(* Logix 5000 project; controller WED2413001_BI600_AB vendor 1 type 14 code 192 rev 35.11; software revision 35.01 *) (continued)
   TRANSITION Tran_008 FROM R00STARTING TO R00EXECUTE
      := EXECUTING
   END_TRANSITION
   STEP R00EXECUTE:
      ACTION Action_008 (N):
         Machine_State:=6;
      END_ACTION
   END_STEP
   TRANSITION Tran_011 FROM R00EXECUTE TO R00STOPPING
      := 
         STOP_CMD
   END_TRANSITION
   TRANSITION Tran_012 FROM R00EXECUTE TO R00COMPLETING
      := PRODUCTION_CNT
   END_TRANSITION
   TRANSITION Tran_009 FROM R00EXECUTE TO R00SUSPENDING
      := SUSPEND_CMD
   END_TRANSITION
   TRANSITION Tran_010 FROM R00EXECUTE TO R00HOLDING
      := HOLD_CMD
   END_TRANSITION
   STEP R00STOPPING:
      ACTION Action_009 (N):
         Machine_State:=7;
      END_ACTION
   END_STEP
   STEP R00COMPLETING:
      ACTION Action_010 (N):
         Machine_State:=16;
      END_ACTION
   END_STEP
   STEP R00SUSPENDING:
      ACTION Action_011 (N):
         Machine_State:=13;
      END_ACTION
   END_STEP
   STEP R00HOLDING:
      ACTION Action_012 (N):
         Machine_State:=10;
      END_ACTION
   END_STEP
   TRANSITION Tran_013 FROM R00STOPPING TO R00STOPPED
      := 1
   END_TRANSITION
   TRANSITION Tran_014 FROM R00COMPLETING TO R00COMPLETE
      := 1
   END_TRANSITION
   TRANSITION Tran_015 FROM R00SUSPENDING TO R00SUSPENDED
      := SUSPEND_CMD
   END_TRANSITION
   TRANSITION Tran_016 FROM R00HOLDING TO R00HELD
      := HOLD_CMD
   END_TRANSITION
   STEP R00COMPLETE:
      ACTION Action_015 (N):
         Machine_State:=17;
      END_ACTION
   END_STEP
   STEP R00SUSPENDED:
      ACTION Action_014 (N):
         Machine_State:=5;
      END_ACTION
   END_STEP
   STEP R00HELD:
      ACTION Action_013 (N):
         Machine_State:=11;
      END_ACTION
   END_STEP
   TRANSITION Tran_017 FROM R00COMPLETE TO R00RESETING
      := 1
   END_TRANSITION
   TRANSITION Tran_018 FROM R00SUSPENDED TO R00UNSUSPENDED
      := SUSPEND_CMD
   END_TRANSITION
   TRANSITION Tran_019 FROM R00HELD TO R00UNHOLDING
      := RESUME_CMD
   END_TRANSITION
   STEP R00UNSUSPENDED:
      ACTION Action_016 (N):
         Machine_State:=14;
      END_ACTION
   END_STEP
   STEP R00UNHOLDING:
      ACTION Action_017 (N):
         Machine_State:=12;
      END_ACTION
   END_STEP
   TRANSITION Tran_020 FROM R00UNSUSPENDED TO R00EXECUTE
      := 1
   END_TRANSITION
   TRANSITION Tran_021 FROM R00UNHOLDING TO R00EXECUTE
      := 1
   END_TRANSITION
END_ROUTINE

ROUTINE R00_Main   (* ladder *)
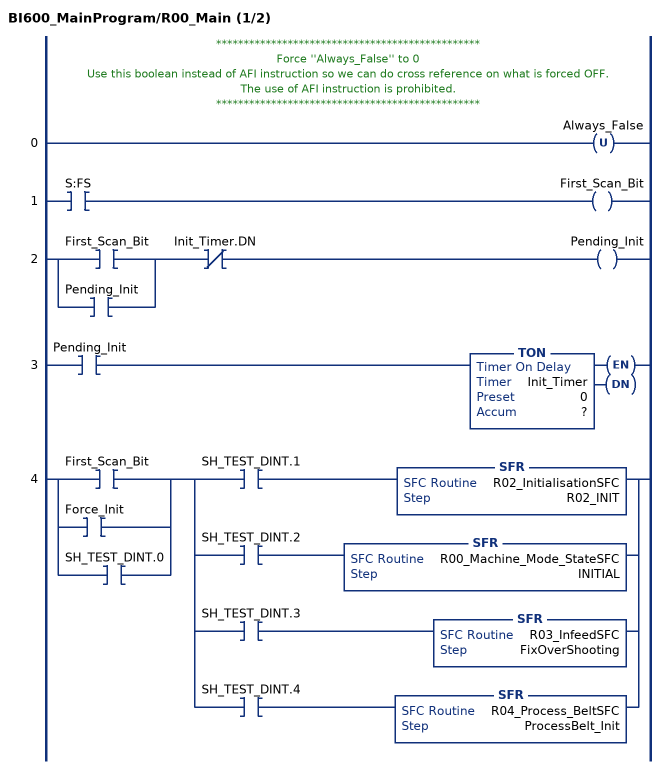
   // ************************************************
   // Force ''Always_False'' to 0
   // Use this boolean instead of AFI instruction so we can do cross reference on what is forced OFF.
   // The use of AFI instruction is prohibited.
   // ************************************************
   0: OTU(Always_False);
   1: XIC(S:FS)OTE(First_Scan_Bit);
   2: [XIC(First_Scan_Bit) ,XIC(Pending_Init) ]XIO(Init_Timer.DN)OTE(Pending_Init);
   3: XIC(Pending_Init)TON(Init_Timer,?,?);
   4: [XIC(First_Scan_Bit) ,XIC(Force_Init) ,XIC(SH_TEST_DINT.0) ][XIC(SH_TEST_DINT.1) SFR(R02_InitialisationSFC,R02_INIT) ,XIC(SH_TEST_DINT.2) SFR(R00_Machine_Mode_StateSFC,INITIAL) ,XIC(SH_TEST_DINT.3) SFR(R03_InfeedSFC,FixOverShooting) ,XIC(SH_TEST_DINT.4) SFR(R04_Process_BeltSFC,ProcessBelt_Init) ];
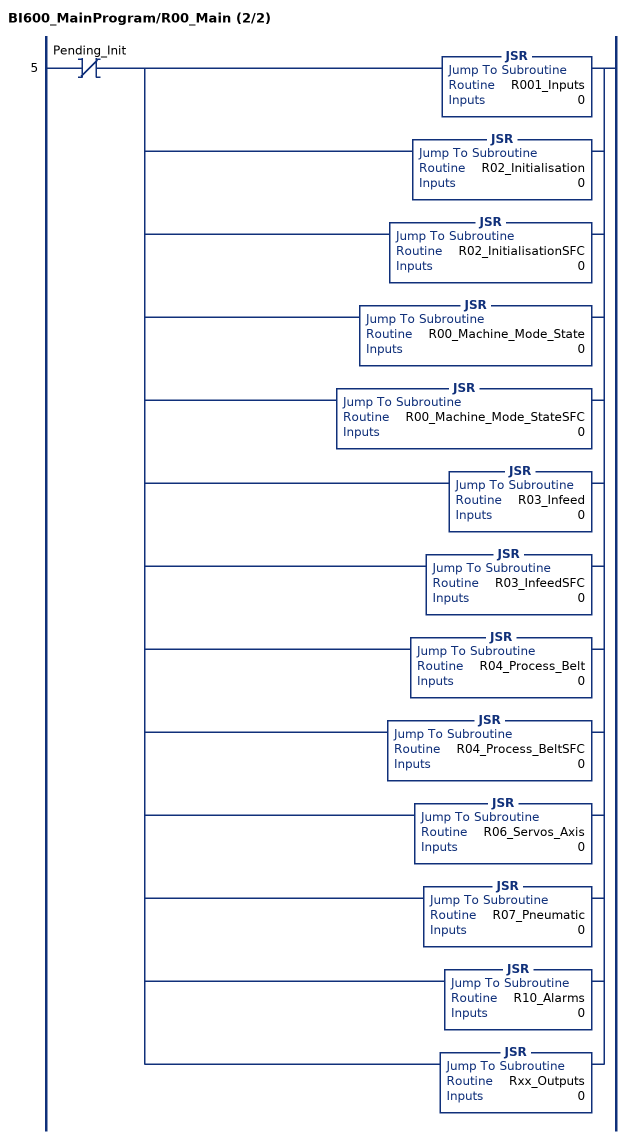
   5: XIO(Pending_Init)[JSR(R001_Inputs,0) ,JSR(R02_Initialisation,0) ,JSR(R02_InitialisationSFC,0) ,JSR(R00_Machine_Mode_State,0) ,JSR(R00_Machine_Mode_StateSFC,0) ,JSR(R03_Infeed,0) ,JSR(R03_InfeedSFC,0) ,JSR(R04_Process_Belt,0) ,JSR(R04_Process_BeltSFC,0) ,JSR(R06_Servos_Axis,0) ,JSR(R07_Pneumatic,0) ,JSR(R10_Alarms,0) ,JSR(Rxx_Outputs,0) ];
END_ROUTINE

ROUTINE R02_Initialisation   (* ladder *)
   // Perform a master reset
   0: NOP();
END_ROUTINE

ROUTINE R02_InitialisationSFC   (* sequential function chart *)
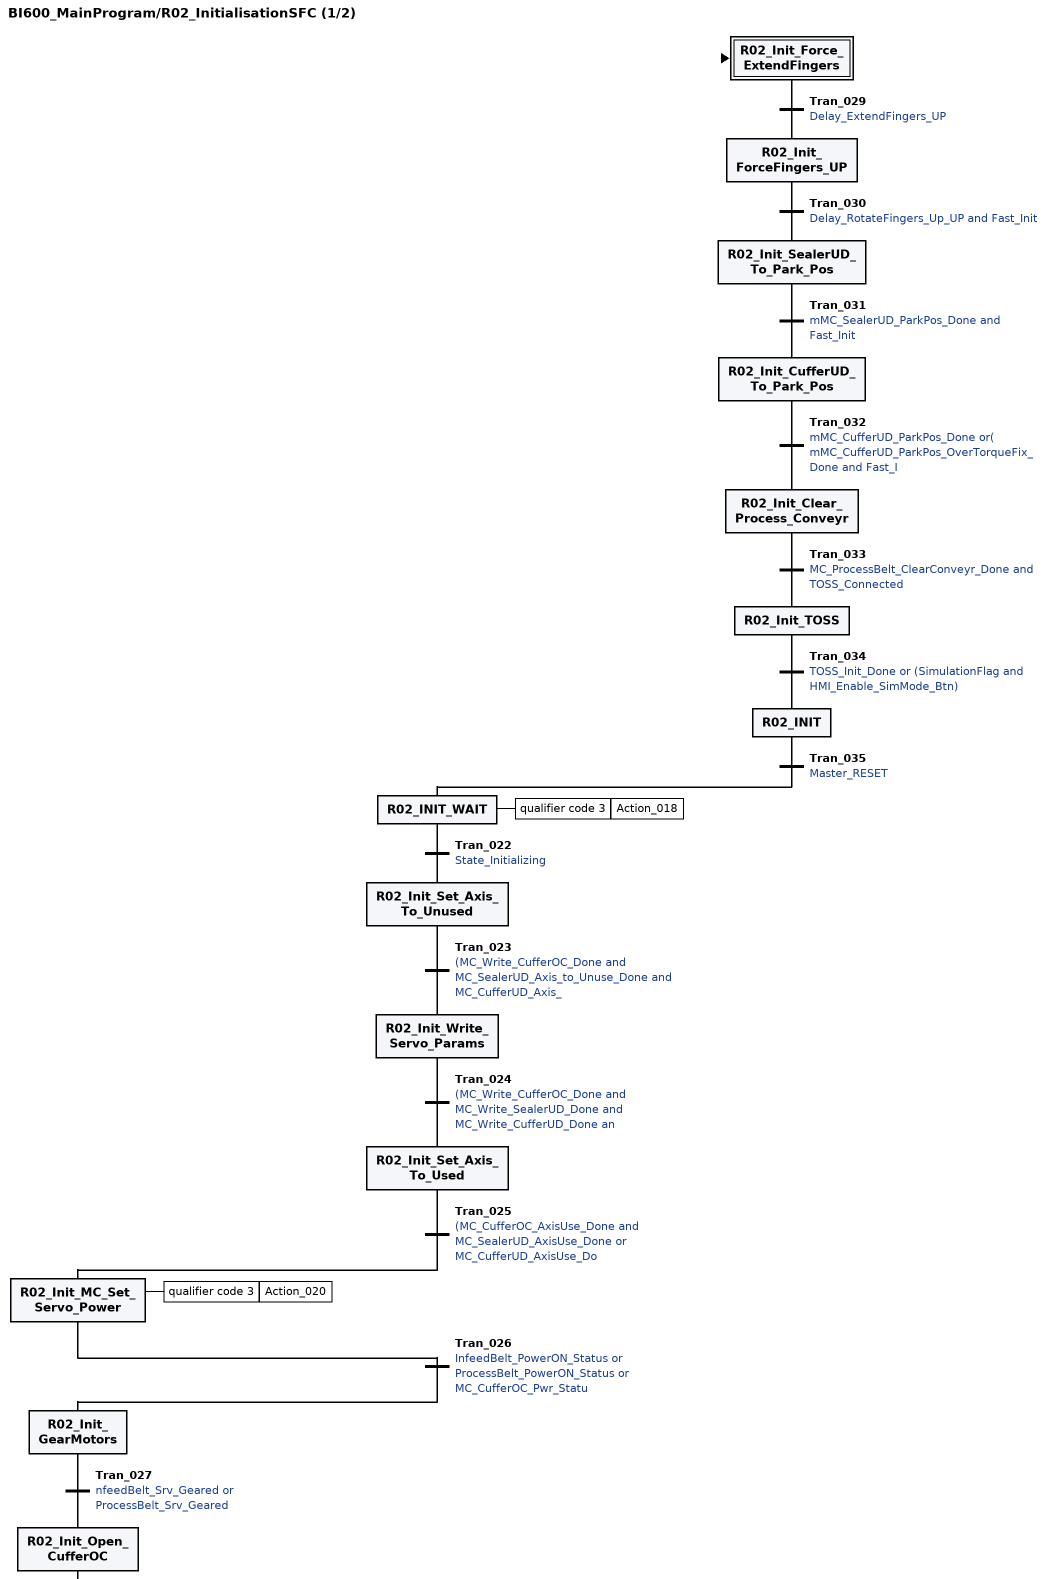
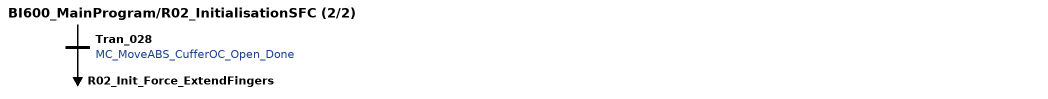
   INITIAL_STEP R02_Init_Force_ExtendFingers:
   END_STEP
   TRANSITION Tran_029 FROM R02_Init_Force_ExtendFingers TO R02_Init_ForceFingers_UP
      := Delay_ExtendFingers_UP
   END_TRANSITION
   STEP R02_INIT_WAIT:
      ACTION Action_018 (qualifier code 3):
         Init_Servo_Power_On :=0;
         Vacuum_ON :=0;
         InfeedBelt_Full_Flag :=0;
         Enable_Full_FilmFeed:=1;
         bBadBagInsert:=0;
      END_ACTION
   END_STEP
   STEP R02_Init_ForceFingers_UP:
   END_STEP
   TRANSITION Tran_022 FROM R02_INIT_WAIT TO R02_Init_Set_Axis_To_Unused
      := State_Initializing
         
   END_TRANSITION
   TRANSITION Tran_030 FROM R02_Init_ForceFingers_UP TO R02_Init_SealerUD_To_Park_Pos
      := Delay_RotateFingers_Up_UP and Fast_Init
   END_TRANSITION
   STEP R02_Init_Set_Axis_To_Unused:
   END_STEP
   STEP R02_Init_SealerUD_To_Park_Pos:
   END_STEP
   TRANSITION Tran_023 FROM R02_Init_Set_Axis_To_Unused TO R02_Init_Write_Servo_Params
      := (MC_Write_CufferOC_Done and
         MC_SealerUD_Axis_to_Unuse_Done and
         MC_CufferUD_Axis_to_Unuse_Done and
         MC_FilmFeed_Axis_to_Unuse_Done and
         mInfeedBelt_MC_AxisToUnuse_Done and
         mProcessBelt_MC_AxisToUnuse_Done) or
         SkipWriteServoPar
   END_TRANSITION
   TRANSITION Tran_031 FROM R02_Init_SealerUD_To_Park_Pos TO R02_Init_CufferUD_To_Park_Pos
      := mMC_SealerUD_ParkPos_Done and Fast_Init
   END_TRANSITION
   STEP R02_Init_Write_Servo_Params:
   END_STEP
   STEP R02_Init_CufferUD_To_Park_Pos:
   END_STEP
   TRANSITION Tran_024 FROM R02_Init_Write_Servo_Params TO R02_Init_Set_Axis_To_Used
      := (MC_Write_CufferOC_Done and
         MC_Write_SealerUD_Done and
         MC_Write_CufferUD_Done and
         MC_Write_FilmFeed_Done and
         mInfeedBelt_MC_WritePar_Done and
         mProcessBelt_MC_WritePar_Done) or
         SkipWriteServoPar
   END_TRANSITION
   TRANSITION Tran_032 FROM R02_Init_CufferUD_To_Park_Pos TO R02_Init_Clear_Process_Conveyr
      := mMC_CufferUD_ParkPos_Done or( mMC_CufferUD_ParkPos_OverTorqueFix_Done and Fast_Init)
   END_TRANSITION
   STEP R02_Init_Set_Axis_To_Used:
   END_STEP
   STEP R02_Init_Clear_Process_Conveyr:
   END_STEP
   TRANSITION Tran_033 FROM R02_Init_Clear_Process_Conveyr TO R02_Init_TOSS
      := MC_ProcessBelt_ClearConveyr_Done and TOSS_Connected
         
   END_TRANSITION
   TRANSITION Tran_025 FROM R02_Init_Set_Axis_To_Used TO R02_Init_MC_Set_Servo_Power
      := (MC_CufferOC_AxisUse_Done and
         MC_SealerUD_AxisUse_Done or
         MC_CufferUD_AxisUse_Done and
         MC_FilmFeed_AxisUse_Done and
         mInfeedBelt_MC_AxisToUse_Done and
         mProcessBelt_MC_AxisToUse_Done)
          or SkipWriteServoPar
   END_TRANSITION
   STEP R02_Init_TOSS:
   END_STEP
   TRANSITION Tran_034 FROM R02_Init_TOSS TO R02_INIT
      := TOSS_Init_Done or (SimulationFlag and HMI_Enable_SimMode_Btn)
   END_TRANSITION
   STEP R02_INIT:
   END_STEP
   STEP R02_Init_MC_Set_Servo_Power:
      ACTION Action_020 (qualifier code 3):
         Init_Servo_Power_On:=1;
      END_ACTION
   END_STEP
   TRANSITION Tran_035 FROM R02_INIT TO R02_INIT_WAIT
      := Master_RESET
   END_TRANSITION
   TRANSITION Tran_026 FROM R02_Init_MC_Set_Servo_Power TO R02_Init_GearMotors
      := InfeedBelt_PowerON_Status or
         ProcessBelt_PowerON_Status or
         MC_CufferOC_Pwr_Status or
         MC_CufferUD_Pwr_Status or
         MC_SealerUD_Pwr_Status or
         MC_FilmFeed_Pwr_Status
   END_TRANSITION
   STEP R02_Init_GearMotors:
   END_STEP
   TRANSITION Tran_027 FROM R02_Init_GearMotors TO R02_Init_Open_CufferOC
      := nfeedBelt_Srv_Geared or ProcessBelt_Srv_Geared
   END_TRANSITION
   STEP R02_Init_Open_CufferOC:
   END_STEP
   TRANSITION Tran_028 FROM R02_Init_Open_CufferOC TO R02_Init_Force_ExtendFingers
      := MC_MoveABS_CufferOC_Open_Done
   END_TRANSITION
END_ROUTINE

ROUTINE R03_Infeed   (* ladder *)
   // Perform a master reset
   0: NOP();
END_ROUTINE

ROUTINE R03_InfeedSFC   (* sequential function chart *)
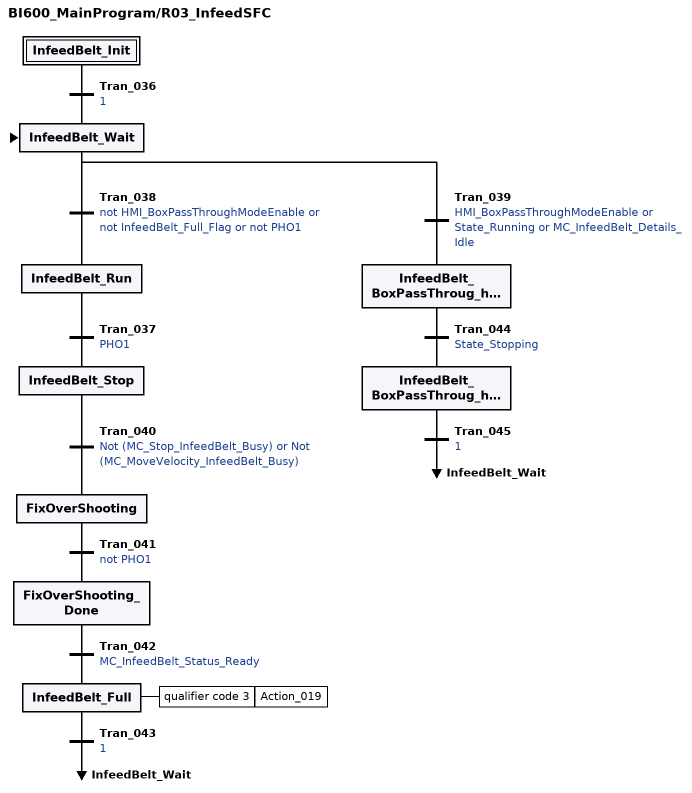
   INITIAL_STEP InfeedBelt_Init:
   END_STEP
   TRANSITION Tran_036 FROM InfeedBelt_Init TO InfeedBelt_Wait
      := 1
   END_TRANSITION
   STEP InfeedBelt_Wait:
   END_STEP
   TRANSITION Tran_038 FROM InfeedBelt_Wait TO InfeedBelt_Run
      := not HMI_BoxPassThroughModeEnable
         or not InfeedBelt_Full_Flag
         or not PHO1
         
         
   END_TRANSITION
   TRANSITION Tran_039 FROM InfeedBelt_Wait TO InfeedBelt_BoxPassThroug_h_Running
      := HMI_BoxPassThroughModeEnable
         or State_Running
         or MC_InfeedBelt_Details_Idle
         
   END_TRANSITION
   STEP InfeedBelt_BoxPassThroug_h_Running:
   END_STEP
   STEP InfeedBelt_Run:
   END_STEP
   TRANSITION Tran_044 FROM InfeedBelt_BoxPassThroug_h_Running TO InfeedBelt_BoxPassThroug_h_Done
      := State_Stopping
         
   END_TRANSITION
   TRANSITION Tran_037 FROM InfeedBelt_Run TO InfeedBelt_Stop
      := PHO1
         
   END_TRANSITION
   STEP InfeedBelt_BoxPassThroug_h_Done:
   END_STEP
   STEP InfeedBelt_Stop:
   END_STEP
   TRANSITION Tran_045 FROM InfeedBelt_BoxPassThroug_h_Done TO InfeedBelt_Wait
      := 1
   END_TRANSITION
   TRANSITION Tran_040 FROM InfeedBelt_Stop TO FixOverShooting
      := Not (MC_Stop_InfeedBelt_Busy) or
         Not (MC_MoveVelocity_InfeedBelt_Busy)
   END_TRANSITION
   STEP FixOverShooting:
   END_STEP
   TRANSITION Tran_041 FROM FixOverShooting TO FixOverShooting_Done
      := not PHO1
         
   END_TRANSITION
   STEP FixOverShooting_Done:
   END_STEP
   TRANSITION Tran_042 FROM FixOverShooting_Done TO InfeedBelt_Full
      := MC_InfeedBelt_Status_Ready
         
   END_TRANSITION
   STEP InfeedBelt_Full:
      ACTION Action_019 (qualifier code 3):
         InfeedBelt_Full_Flag:=1;
      END_ACTION
   END_STEP
   TRANSITION Tran_043 FROM InfeedBelt_Full TO InfeedBelt_Wait
      := 1
   END_TRANSITION
END_ROUTINE

ROUTINE R04_Process_Belt   (* ladder *)
   0: NOP();
END_ROUTINE

ROUTINE R04_Process_BeltSFC   (* sequential function chart *)
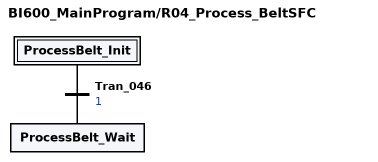
   INITIAL_STEP ProcessBelt_Init:
   END_STEP
   TRANSITION Tran_046 FROM ProcessBelt_Init TO ProcessBelt_Wait
      := 1
   END_TRANSITION
   STEP ProcessBelt_Wait:
   END_STEP
END_ROUTINE

ROUTINE R06_Servos_Axis   (* ladder *)
   0: NOP();
END_ROUTINE

ROUTINE R07_Pneumatic   (* ladder *)
   0: NOP();
END_ROUTINE

ROUTINE R10_Alarms   (* ladder *)
   0: NOP();
END_ROUTINE

ROUTINE Rxx_Outputs   (* ladder *)
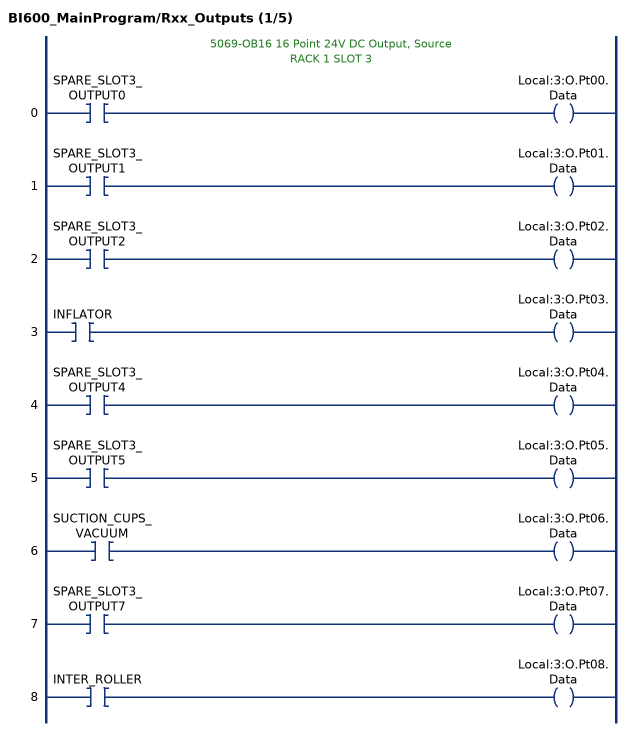
   // 5069-OB16 16 Point 24V DC Output, Source
   // RACK 1 SLOT 3
   0: XIC(SPARE_SLOT3_OUTPUT0)OTE(Local:3:O.Pt00.Data);
   1: XIC(SPARE_SLOT3_OUTPUT1)OTE(Local:3:O.Pt01.Data);
   2: XIC(SPARE_SLOT3_OUTPUT2)OTE(Local:3:O.Pt02.Data);
   3: XIC(INFLATOR)OTE(Local:3:O.Pt03.Data);
   4: XIC(SPARE_SLOT3_OUTPUT4)OTE(Local:3:O.Pt04.Data);
   5: XIC(SPARE_SLOT3_OUTPUT5)OTE(Local:3:O.Pt05.Data);
   6: XIC(SUCTION_CUPS_VACUUM)OTE(Local:3:O.Pt06.Data);
   7: XIC(SPARE_SLOT3_OUTPUT7)OTE(Local:3:O.Pt07.Data);
   8: XIC(INTER_ROLLER)OTE(Local:3:O.Pt08.Data);
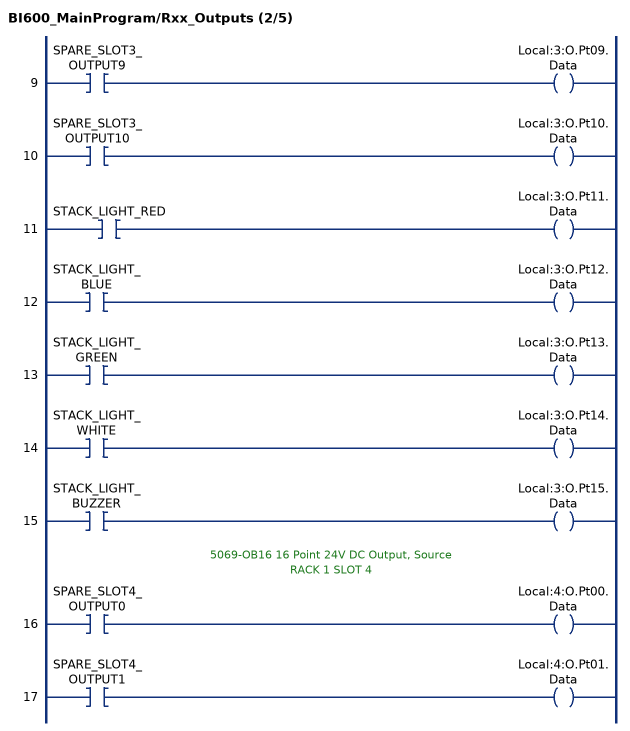
   9: XIC(SPARE_SLOT3_OUTPUT9)OTE(Local:3:O.Pt09.Data);
   10: XIC(SPARE_SLOT3_OUTPUT10)OTE(Local:3:O.Pt10.Data);
   11: XIC(STACK_LIGHT_RED)OTE(Local:3:O.Pt11.Data);
   12: XIC(STACK_LIGHT_BLUE)OTE(Local:3:O.Pt12.Data);
   13: XIC(STACK_LIGHT_GREEN)OTE(Local:3:O.Pt13.Data);
   14: XIC(STACK_LIGHT_WHITE)OTE(Local:3:O.Pt14.Data);
   15: XIC(STACK_LIGHT_BUZZER)OTE(Local:3:O.Pt15.Data);
   // 5069-OB16 16 Point 24V DC Output, Source
   // RACK 1 SLOT 4
   16: XIC(SPARE_SLOT4_OUTPUT0)OTE(Local:4:O.Pt00.Data);
   17: XIC(SPARE_SLOT4_OUTPUT1)OTE(Local:4:O.Pt01.Data);
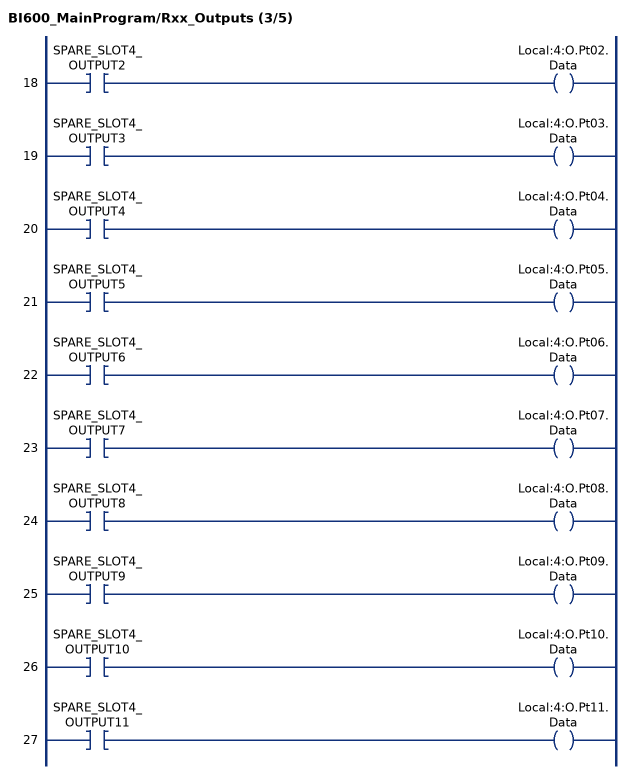
   18: XIC(SPARE_SLOT4_OUTPUT2)OTE(Local:4:O.Pt02.Data);
   19: XIC(SPARE_SLOT4_OUTPUT3)OTE(Local:4:O.Pt03.Data);
   20: XIC(SPARE_SLOT4_OUTPUT4)OTE(Local:4:O.Pt04.Data);
   21: XIC(SPARE_SLOT4_OUTPUT5)OTE(Local:4:O.Pt05.Data);
   22: XIC(SPARE_SLOT4_OUTPUT6)OTE(Local:4:O.Pt06.Data);
   23: XIC(SPARE_SLOT4_OUTPUT7)OTE(Local:4:O.Pt07.Data);
   24: XIC(SPARE_SLOT4_OUTPUT8)OTE(Local:4:O.Pt08.Data);
   25: XIC(SPARE_SLOT4_OUTPUT9)OTE(Local:4:O.Pt09.Data);
   26: XIC(SPARE_SLOT4_OUTPUT10)OTE(Local:4:O.Pt10.Data);
   27: XIC(SPARE_SLOT4_OUTPUT11)OTE(Local:4:O.Pt11.Data);
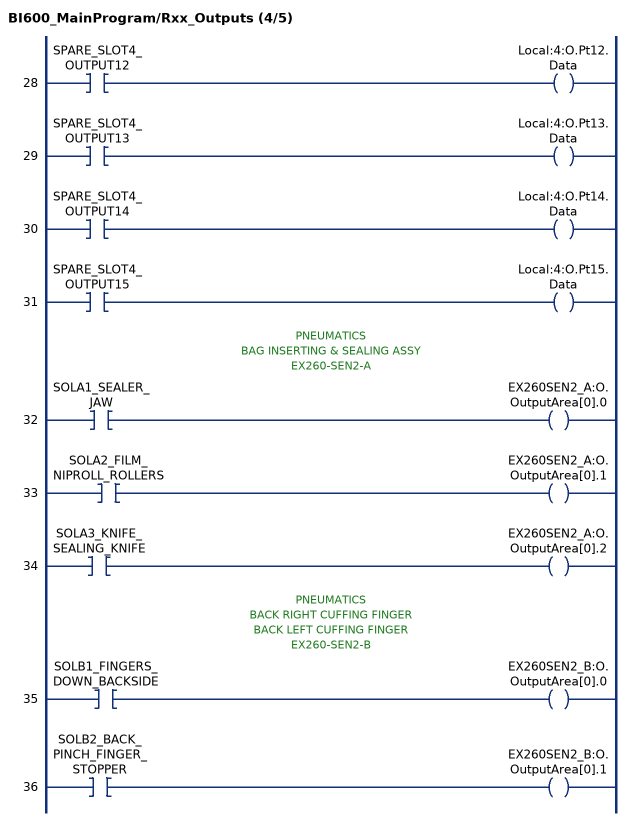
   28: XIC(SPARE_SLOT4_OUTPUT12)OTE(Local:4:O.Pt12.Data);
   29: XIC(SPARE_SLOT4_OUTPUT13)OTE(Local:4:O.Pt13.Data);
   30: XIC(SPARE_SLOT4_OUTPUT14)OTE(Local:4:O.Pt14.Data);
   31: XIC(SPARE_SLOT4_OUTPUT15)OTE(Local:4:O.Pt15.Data);
   // PNEUMATICS
   // BAG INSERTING & SEALING ASSY
   // EX260-SEN2-A
   32: XIC(SOLA1_SEALER_JAW)OTE(EX260SEN2_A:O.OutputArea[0].0);
   33: XIC(SOLA2_FILM_NIPROLL_ROLLERS)OTE(EX260SEN2_A:O.OutputArea[0].1);
   34: XIC(SOLA3_KNIFE_SEALING_KNIFE)OTE(EX260SEN2_A:O.OutputArea[0].2);
   // PNEUMATICS
   // BACK RIGHT CUFFING FINGER
   // BACK LEFT CUFFING FINGER
   // EX260-SEN2-B
   35: XIC(SOLB1_FINGERS_DOWN_BACKSIDE)OTE(EX260SEN2_B:O.OutputArea[0].0);
   36: XIC(SOLB2_BACK_PINCH_FINGER_STOPPER)OTE(EX260SEN2_B:O.OutputArea[0].1);
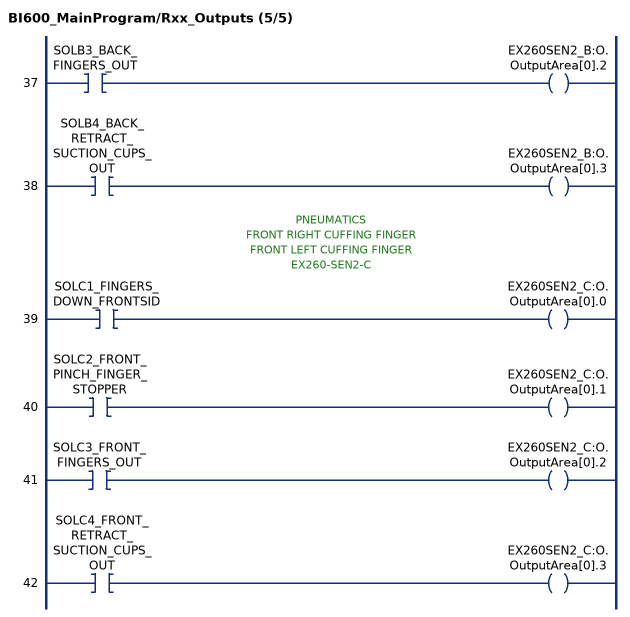
   37: XIC(SOLB3_BACK_FINGERS_OUT)OTE(EX260SEN2_B:O.OutputArea[0].2);
   38: XIC(SOLB4_BACK_RETRACT_SUCTION_CUPS_OUT)OTE(EX260SEN2_B:O.OutputArea[0].3);
   // PNEUMATICS
   // FRONT RIGHT CUFFING FINGER
   // FRONT LEFT CUFFING FINGER
   // EX260-SEN2-C
   39: XIC(SOLC1_FINGERS_DOWN_FRONTSID)OTE(EX260SEN2_C:O.OutputArea[0].0);
   40: XIC(SOLC2_FRONT_PINCH_FINGER_STOPPER)OTE(EX260SEN2_C:O.OutputArea[0].1);
   41: XIC(SOLC3_FRONT_FINGERS_OUT)OTE(EX260SEN2_C:O.OutputArea[0].2);
   42: XIC(SOLC4_FRONT_RETRACT_SUCTION_CUPS_OUT)OTE(EX260SEN2_C:O.OutputArea[0].3);
END_ROUTINE
END_PROGRAM
